REGION Network 14: Reset Manual Mode
   // Reset Manual mode when loose input flag of manual orremote enable kicks in
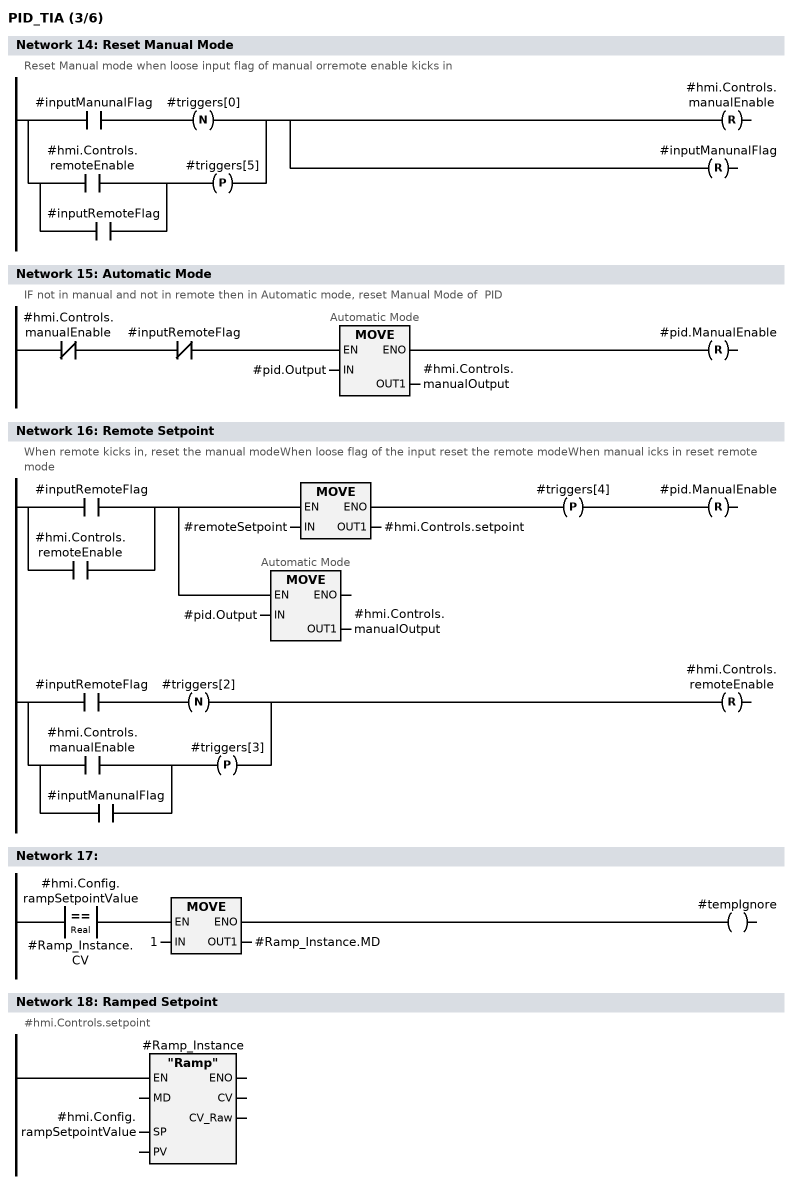
   RUNG wire#powerrail
      Contact( #inputManunalFlag )
      N_Trig( #triggers[0] )
      wire#w1
      R_Coil( #hmi.Controls.manualEnable )
   END_RUNG
   RUNG wire#powerrail
      Contact( #hmi.Controls.remoteEnable )
      wire#w2
      P_Trig( #triggers[5] )
   END_RUNG wire#w1
   RUNG wire#powerrail
      Contact( #inputRemoteFlag )
   END_RUNG wire#w2
   RUNG wire#w1
      R_Coil( #inputManunalFlag )
   END_RUNG
   // the same network as SCL:
   #_w1 := NOT #inputManunalFlag AND #triggers[0];   // falling edge
   #triggers[0] := #inputManunalFlag;
   #_w2 := #hmi.Controls.remoteEnable OR #inputRemoteFlag;
   #_w3 := #_w2 AND NOT #triggers[5];   // rising edge
   #triggers[5] := #_w2;
   IF #_w1 OR #_w3 THEN
       #hmi.Controls.manualEnable := FALSE;
       #inputManunalFlag := FALSE;
   END_IF;
END_REGION

REGION Network 15: Automatic Mode
   // IF not in manual and not in remote then in Automatic mode, reset Manual Mode of  PID
   RUNG wire#powerrail
      I_Contact( #hmi.Controls.manualEnable )
      I_Contact( #inputRemoteFlag )
      Move(in := #pid.Output, out1 => #hmi.Controls.manualOutput)   // Automatic Mode
      R_Coil( #pid.ManualEnable )
   END_RUNG
   // the same network as SCL:
   IF NOT #hmi.Controls.manualEnable AND NOT #inputRemoteFlag THEN
       #hmi.Controls.manualOutput := #pid.Output;   // Automatic Mode
       #pid.ManualEnable := FALSE;
   END_IF;
END_REGION

REGION Network 16: Remote Setpoint
   // When remote kicks in, reset the manual modeWhen loose flag of the input reset the remote modeWhen manual icks in reset remote mode
   RUNG wire#powerrail
      Contact( #inputRemoteFlag )
      wire#w1
      Move(in := #remoteSetpoint, out1 => #hmi.Controls.setpoint)
      P_Trig( #triggers[4] )
      R_Coil( #pid.ManualEnable )
   END_RUNG
   RUNG wire#powerrail
      Contact( #hmi.Controls.remoteEnable )
   END_RUNG wire#w1
   RUNG wire#w1
      Move(in := #pid.Output, out1 => #hmi.Controls.manualOutput)   // Automatic Mode
   END_RUNG
   RUNG wire#powerrail
      Contact( #inputRemoteFlag )
      N_Trig( #triggers[2] )
      wire#w2
      R_Coil( #hmi.Controls.remoteEnable )
   END_RUNG
   RUNG wire#powerrail
      Contact( #hmi.Controls.manualEnable )
      wire#w3
      P_Trig( #triggers[3] )
   END_RUNG wire#w2
   RUNG wire#powerrail
      Contact( #inputManunalFlag )
   END_RUNG wire#w3
   // the same network as SCL:
   #_w1 := #inputRemoteFlag OR #hmi.Controls.remoteEnable;
   IF #_w1 THEN #hmi.Controls.setpoint := #remoteSetpoint; END_IF;
   #_w2 := #_w1 AND NOT #triggers[4];   // rising edge
   #triggers[4] := #_w1;
   IF #_w2 THEN #pid.ManualEnable := FALSE; END_IF;
   IF #_w1 THEN
       #hmi.Controls.manualOutput := #pid.Output;   // Automatic Mode
   END_IF;
   #_w3 := NOT #inputRemoteFlag AND #triggers[2];   // falling edge
   #triggers[2] := #inputRemoteFlag;
   #_w4 := #hmi.Controls.manualEnable OR #inputManunalFlag;
   #_w5 := #_w4 AND NOT #triggers[3];   // rising edge
   #triggers[3] := #_w4;
   IF #_w3 OR #_w5 THEN #hmi.Controls.remoteEnable := FALSE; END_IF;
END_REGION

REGION Network 17
   RUNG wire#powerrail
      { S7_Templates := "SrcType := Real" } EQ_Contact(in1 := #hmi.Config.rampSetpointValue, in2 := #Ramp_Instance.CV)
      Move(in := 1, out1 => #Ramp_Instance.MD)
      Coil( #tempIgnore )
   END_RUNG
   // the same network as SCL:
   #_w1 := #hmi.Config.rampSetpointValue = #Ramp_Instance.CV;
   IF #_w1 THEN #Ramp_Instance.MD := 1; END_IF;
   #tempIgnore := #_w1;
END_REGION

REGION Network 18: Ramped Setpoint
   // #hmi.Controls.setpoint
   RUNG wire#powerrail
      #Ramp_Instance(MD :=, SP := #hmi.Config.rampSetpointValue, PV :=, CV =>, CV_Raw =>)
   END_RUNG
   // the same network as SCL:
   #Ramp_Instance(SP := #hmi.Config.rampSetpointValue);   // "Ramp"
END_REGION

REGION Network 19: Setpoint Control
   // If ramp enabled then move ramped setpointif ramp disabled then move hmi setpoint
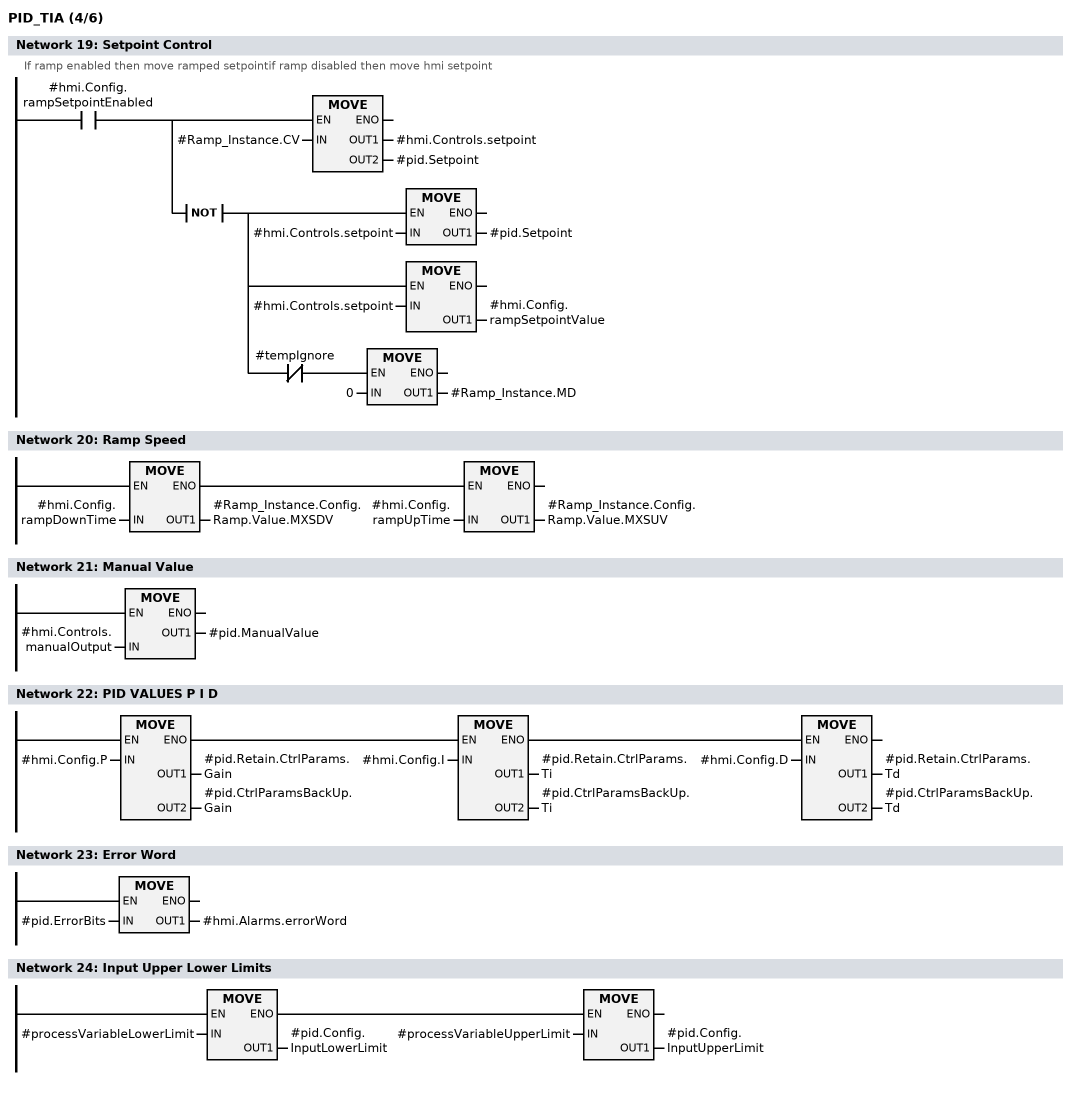
   RUNG wire#powerrail
      Contact( #hmi.Config.rampSetpointEnabled )
      wire#w1
      Move(in := #Ramp_Instance.CV, out1 => #hmi.Controls.setpoint, out2 => #pid.Setpoint)
   END_RUNG
   RUNG wire#w1
      Not()
      wire#w2
      Move(in := #hmi.Controls.setpoint, out1 => #pid.Setpoint)
   END_RUNG
   RUNG wire#w2
      Move(in := #hmi.Controls.setpoint, out1 => #hmi.Config.rampSetpointValue)
   END_RUNG
   RUNG wire#w2
      I_Contact( #tempIgnore )
      Move(in := 0, out1 => #Ramp_Instance.MD)
   END_RUNG
   // the same network as SCL:
   IF #hmi.Config.rampSetpointEnabled THEN
       #hmi.Controls.setpoint := #Ramp_Instance.CV;
       #pid.Setpoint := #Ramp_Instance.CV;
   END_IF;
   #_w1 := NOT #hmi.Config.rampSetpointEnabled;
   IF #_w1 THEN
       #pid.Setpoint := #hmi.Controls.setpoint;
       #hmi.Config.rampSetpointValue := #hmi.Controls.setpoint;
   END_IF;
   IF #_w1 AND NOT #tempIgnore THEN #Ramp_Instance.MD := 0; END_IF;
END_REGION

REGION Network 20: Ramp Speed
   RUNG wire#powerrail
      Move(in := #hmi.Config.rampDownTime, out1 => #Ramp_Instance.Config.Ramp.Value.MXSDV)
      Move(in := #hmi.Config.rampUpTime, out1 => #Ramp_Instance.Config.Ramp.Value.MXSUV)
   END_RUNG
   // the same network as SCL:
   #Ramp_Instance.Config.Ramp.Value.MXSDV := #hmi.Config.rampDownTime;
   #Ramp_Instance.Config.Ramp.Value.MXSUV := #hmi.Config.rampUpTime;
END_REGION

REGION Network 21: Manual Value
   RUNG wire#powerrail
      Move(in := #hmi.Controls.manualOutput, out1 => #pid.ManualValue)
   END_RUNG
   // the same network as SCL:
   #pid.ManualValue := #hmi.Controls.manualOutput;
END_REGION

REGION Network 22: PID VALUES P I D
   RUNG wire#powerrail
      Move(in := #hmi.Config.P, out1 => #pid.Retain.CtrlParams.Gain, out2 => #pid.CtrlParamsBackUp.Gain)
      Move(in := #hmi.Config.I, out1 => #pid.Retain.CtrlParams.Ti, out2 => #pid.CtrlParamsBackUp.Ti)
      Move(in := #hmi.Config.D, out1 => #pid.Retain.CtrlParams.Td, out2 => #pid.CtrlParamsBackUp.Td)
   END_RUNG
   // the same network as SCL:
   #pid.Retain.CtrlParams.Gain := #hmi.Config.P;
   #pid.CtrlParamsBackUp.Gain := #hmi.Config.P;
   #pid.Retain.CtrlParams.Ti := #hmi.Config.I;
   #pid.CtrlParamsBackUp.Ti := #hmi.Config.I;
   #pid.Retain.CtrlParams.Td := #hmi.Config.D;
   #pid.CtrlParamsBackUp.Td := #hmi.Config.D;
END_REGION

REGION Network 23: Error Word
   RUNG wire#powerrail
      Move(in := #pid.ErrorBits, out1 => #hmi.Alarms.errorWord)
   END_RUNG
   // the same network as SCL:
   #hmi.Alarms.errorWord := #pid.ErrorBits;
END_REGION

REGION Network 24: Input Upper Lower Limits
   RUNG wire#powerrail
      Move(in := #processVariableLowerLimit, out1 => #pid.Config.InputLowerLimit)
      Move(in := #processVariableUpperLimit, out1 => #pid.Config.InputUpperLimit)
   END_RUNG
   // the same network as SCL:
   #pid.Config.InputLowerLimit := #processVariableLowerLimit;
   #pid.Config.InputUpperLimit := #processVariableUpperLimit;
END_REGION

REGION Network 25: Input to Input PID
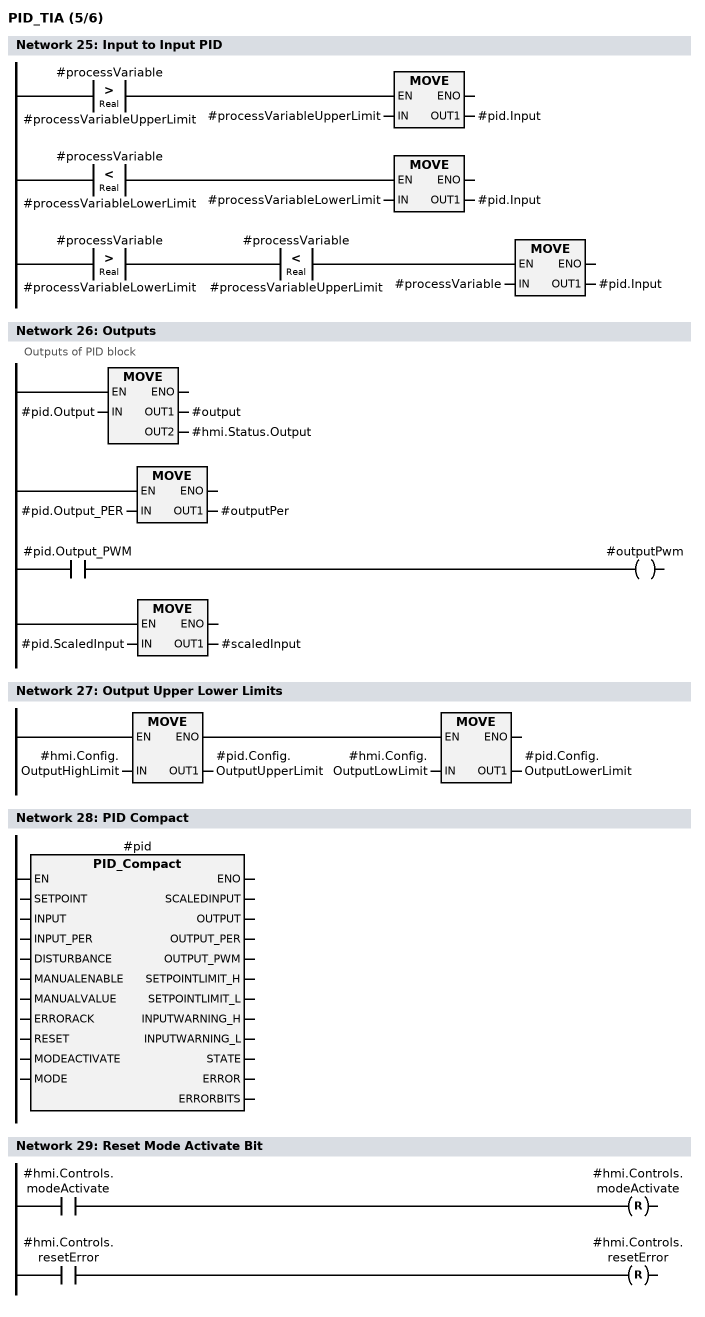
   RUNG wire#powerrail
      { S7_Templates := "SrcType := Real" } GT_Contact(in1 := #processVariable, in2 := #processVariableUpperLimit)
      Move(in := #processVariableUpperLimit, out1 => #pid.Input)
   END_RUNG
   RUNG wire#powerrail
      { S7_Templates := "SrcType := Real" } LT_Contact(in1 := #processVariable, in2 := #processVariableLowerLimit)
      Move(in := #processVariableLowerLimit, out1 => #pid.Input)
   END_RUNG
   RUNG wire#powerrail
      { S7_Templates := "SrcType := Real" } GT_Contact(in1 := #processVariable, in2 := #processVariableLowerLimit)
      { S7_Templates := "SrcType := Real" } LT_Contact(in1 := #processVariable, in2 := #processVariableUpperLimit)
      Move(in := #processVariable, out1 => #pid.Input)
   END_RUNG
   // the same network as SCL:
   IF #processVariable > #processVariableUpperLimit THEN #pid.Input := #processVariableUpperLimit; END_IF;
   IF #processVariable < #processVariableLowerLimit THEN #pid.Input := #processVariableLowerLimit; END_IF;
   IF (#processVariable > #processVariableLowerLimit) AND (#processVariable < #processVariableUpperLimit) THEN
       #pid.Input := #processVariable;
   END_IF;
END_REGION

REGION Network 26: Outputs
   // Outputs of PID block
   RUNG wire#powerrail
      Move(in := #pid.Output, out1 => #output, out2 => #hmi.Status.Output)
   END_RUNG
   RUNG wire#powerrail
      Move(in := #pid.Output_PER, out1 => #outputPer)
   END_RUNG
   RUNG wire#powerrail
      Contact( #pid.Output_PWM )
      Coil( #outputPwm )
   END_RUNG
   RUNG wire#powerrail
      Move(in := #pid.ScaledInput, out1 => #scaledInput)
   END_RUNG
   // the same network as SCL:
   #output := #pid.Output;
   #hmi.Status.Output := #pid.Output;
   #outputPer := #pid.Output_PER;
   #outputPwm := #pid.Output_PWM;
   #scaledInput := #pid.ScaledInput;
END_REGION

REGION Network 27: Output Upper Lower Limits
   RUNG wire#powerrail
      Move(in := #hmi.Config.OutputHighLimit, out1 => #pid.Config.OutputUpperLimit)
      Move(in := #hmi.Config.OutputLowLimit, out1 => #pid.Config.OutputLowerLimit)
   END_RUNG
   // the same network as SCL:
   #pid.Config.OutputUpperLimit := #hmi.Config.OutputHighLimit;
   #pid.Config.OutputLowerLimit := #hmi.Config.OutputLowLimit;
END_REGION

REGION Network 28: PID Compact
   #pid();   // PID_Compact
END_REGION

REGION Network 29: Reset Mode Activate Bit
   RUNG wire#powerrail
      Contact( #hmi.Controls.modeActivate )
      R_Coil( #hmi.Controls.modeActivate )
   END_RUNG
   RUNG wire#powerrail
      Contact( #hmi.Controls.resetError )
      R_Coil( #hmi.Controls.resetError )
   END_RUNG
   // the same network as SCL:
   IF #hmi.Controls.modeActivate THEN #hmi.Controls.modeActivate := FALSE; END_IF;
   IF #hmi.Controls.resetError THEN #hmi.Controls.resetError := FALSE; END_IF;
END_REGION

REGION Network 30: PV Tracking
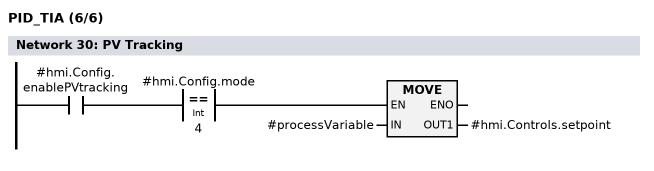
   RUNG wire#powerrail
      Contact( #hmi.Config.enablePVtracking )
      { S7_Templates := "SrcType := Int" } EQ_Contact(in1 := #hmi.Config.mode, in2 := 4)
      Move(in := #processVariable, out1 => #hmi.Controls.setpoint)
   END_RUNG
   // the same network as SCL:
   IF #hmi.Config.enablePVtracking AND (#hmi.Config.mode = 4) THEN
       #hmi.Controls.setpoint := #processVariable;
   END_IF;
END_REGION
END_FUNCTION_BLOCK

// folder: 1}Library/Pumps

FUNCTION_BLOCK "SimpleMotorStater"   // FB823, LAD
{ S7_Optimized_Access := 'TRUE' }
VERSION : 0.1
   VAR_INPUT
      OP_Mode : Bool;   // Output Mode for the Stop CMD if True( Normal Open Output) If False ( Normal Close Output)
      ON : Bool;   // Motor On
      OFF : Bool := TRUE;   // Motor OFF
      CF : Bool;   // Status- Contact Feedback
      IL : Bool := TRUE;   // status-Interlock
      "Lead Control" : Bool := TRUE;
   END_VAR
   VAR_OUTPUT
      Stop_CMD : Bool := TRUE;   // Stop Command for the Motor
      Start_CMD : Bool;   // Start Command for the Motor
      RST : Bool;   // Reset Overload
   END_VAR
   VAR
      HMI : Struct   // Data Struct for HMI
         Controls : Struct
            Start : Bool;
            Stop : Bool := TRUE;
            Reset : Bool;
            Lockout : Bool;
         END_STRUCT;
         Status : Struct
            Mode : Bool;   // Output Mode for the Stop CMD if True Normal Open Output (NO) If False Normal Close Output (NC)
            CF : Bool;   // Status- Contact Feedback
            IL : Bool;   // Status-Interlock
            State : Int;   // 0=off, 1=on, 2=fault,3= Lockout
         END_STRUCT;
      END_STRUCT;
   END_VAR
   VAR RETAIN
      Config : Struct
         HMI : Struct
            Start_PT : Time := T#500MS;   // Start CMD Pulse Time
            Stop_PT : Time := T#500MS;   // Stop CMD Pulse Time
            CF_Delay : Time := T#10s;   // Contact Feedback Delay Time
            NCresetDelay : Time := T#1s;   // time to Set stop on went in NC Mode
            Enable_HMI_Controls : Int;   // MODE 1 PLC CTRL / MODE 2 HMII
         END_STRUCT;
      END_STRUCT;
   END_VAR
   VAR
      OS : Struct
         ON : Bool;
         OFF : Bool;
         HMION : Bool;
         HMIOFF : Bool;
         CF_PULSE : Bool;
         ILPOS : Bool;
         PULSE : Bool;
      END_STRUCT;
      STOP_CMD_TOF : TOF_TIME;   // Stop CMD Pulse Timer
      START_CMD_TOF : TOF_TIME;   // Start CMD Pulse Timer
      CF_Delay_TON : TOF_TIME;   // Contact Feedback Delay Timer
      DelayforReset : TON_TIME;
      FaultTimer : IEC_TIMER;
      Fault : Bool;
      "Lockout Trig" : Bool;
   END_VAR
   VAR_TEMP
      STOP : Bool;
   END_VAR
   VAR_TEMP   // added for the SCL form of the ladder/FBD networks
      _w1 : Bool;
      _w2 : Bool;
      _w3 : Bool;
      _w4 : Bool;
      _w5 : Bool;
      _w6 : Bool;
      _w7 : Bool;
      _w8 : Bool;
   END_VAR
BEGIN

REGION Network 1: Status-Interlock
   // Interloack Status for HMI
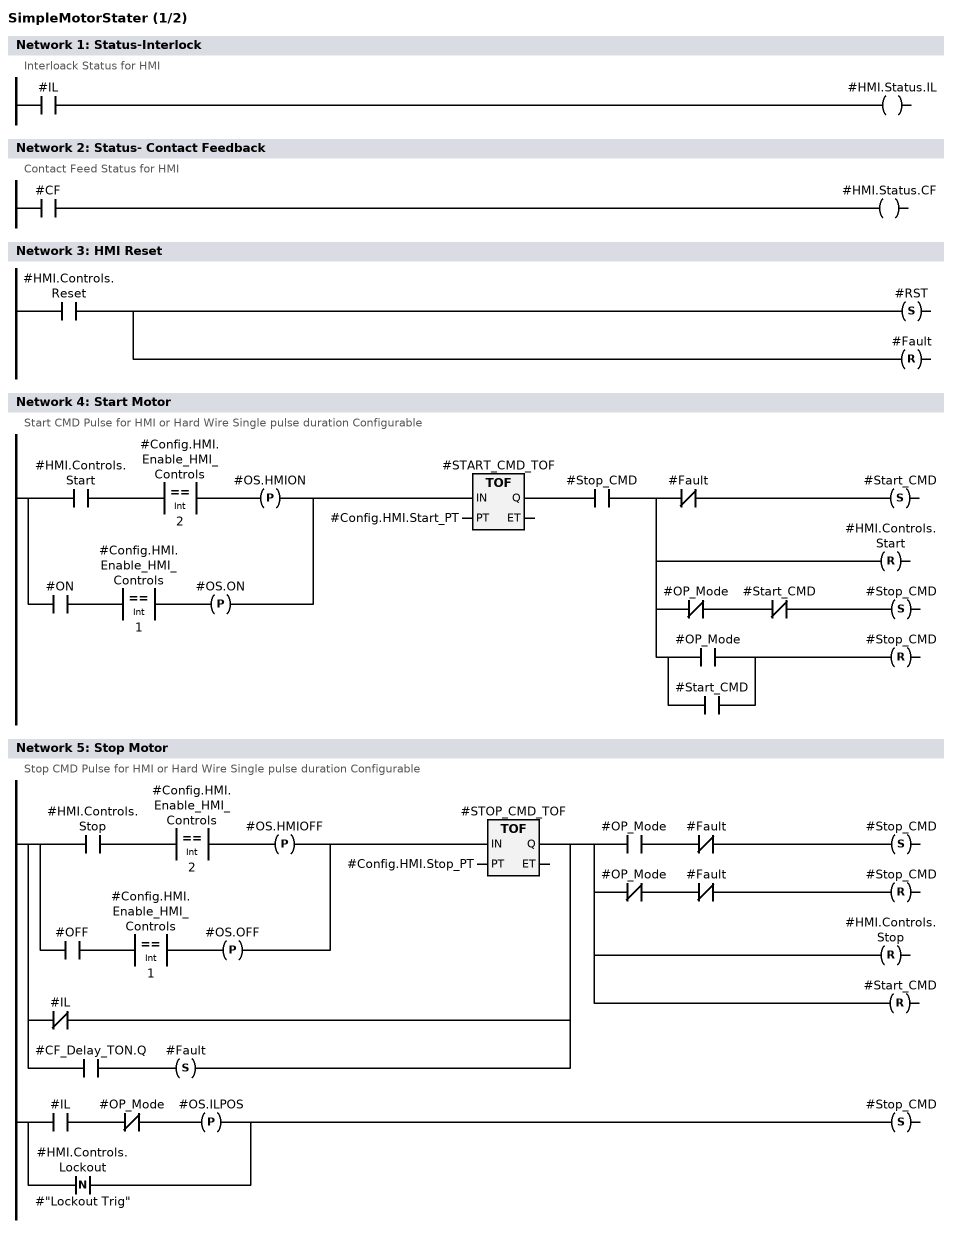
   RUNG wire#powerrail
      Contact( #IL )
      Coil( #HMI.Status.IL )
   END_RUNG
   // the same network as SCL:
   #HMI.Status.IL := #IL;
END_REGION

REGION Network 2: Status- Contact Feedback
   // Contact Feed Status for HMI
   RUNG wire#powerrail
      Contact( #CF )
      Coil( #HMI.Status.CF )
   END_RUNG
   // the same network as SCL:
   #HMI.Status.CF := #CF;
END_REGION

REGION Network 3: HMI Reset
   RUNG wire#powerrail
      Contact( #HMI.Controls.Reset )
      wire#w1
      S_Coil( #RST )
   END_RUNG
   RUNG wire#w1
      R_Coil( #Fault )
   END_RUNG
   // the same network as SCL:
   IF #HMI.Controls.Reset THEN
       #RST := TRUE;
       #Fault := FALSE;
   END_IF;
END_REGION

REGION Network 4: Start Motor
   // Start CMD Pulse for HMI or Hard Wire Single pulse duration Configurable
   #_w1 := #HMI.Controls.Start AND (#Config.HMI.Enable_HMI_Controls = 2);
   #_w2 := #_w1 AND NOT #OS.HMION;   // rising edge
   #OS.HMION := #_w1;
   #_w3 := #ON AND (#Config.HMI.Enable_HMI_Controls = 1);
   #_w4 := #_w3 AND NOT #OS.ON;   // rising edge
   #OS.ON := #_w3;
   #START_CMD_TOF(IN := #_w2 OR #_w4, PT := #Config.HMI.Start_PT);   // TOF
   #_w5 := #START_CMD_TOF.Q AND #Stop_CMD;
   IF #_w5 AND NOT #Fault THEN #Start_CMD := TRUE; END_IF;
   IF #_w5 THEN #HMI.Controls.Start := FALSE; END_IF;
   IF #_w5 AND NOT #OP_Mode AND NOT #Start_CMD THEN #Stop_CMD := TRUE; END_IF;
   IF #_w5 AND (#OP_Mode OR #Start_CMD) THEN #Stop_CMD := FALSE; END_IF;
END_REGION

REGION Network 5: Stop Motor
   // Stop CMD Pulse for HMI or Hard Wire Single pulse duration Configurable
   #_w1 := #HMI.Controls.Stop AND (#Config.HMI.Enable_HMI_Controls = 2);
   #_w2 := #_w1 AND NOT #OS.HMIOFF;   // rising edge
   #OS.HMIOFF := #_w1;
   #_w3 := #OFF AND (#Config.HMI.Enable_HMI_Controls = 1);
   #_w4 := #_w3 AND NOT #OS.OFF;   // rising edge
   #OS.OFF := #_w3;
   #STOP_CMD_TOF(IN := #_w2 OR #_w4, PT := #Config.HMI.Stop_PT);   // TOF
   IF #CF_Delay_TON.Q THEN #Fault := TRUE; END_IF;
   #_w5 := #STOP_CMD_TOF.Q OR NOT #IL OR #CF_Delay_TON.Q;
   IF #_w5 AND #OP_Mode AND NOT #Fault THEN #Stop_CMD := TRUE; END_IF;
   IF #_w5 AND NOT #OP_Mode AND NOT #Fault THEN #Stop_CMD := FALSE; END_IF;
   IF #_w5 THEN
       #HMI.Controls.Stop := FALSE;
       #Start_CMD := FALSE;
   END_IF;
   #_w6 := #IL AND NOT #OP_Mode;
   #_w7 := #_w6 AND NOT #OS.ILPOS;   // rising edge
   #OS.ILPOS := #_w6;
   #_w8 := NOT #HMI.Controls.Lockout AND #"Lockout Trig";   // falling edge of #HMI.Controls.Lockout
   #"Lockout Trig" := #HMI.Controls.Lockout;
   IF #_w7 OR #_w8 THEN #Stop_CMD := TRUE; END_IF;
END_REGION

REGION Network 6: Delay for Contact feedback
   // Timer Delay for For Feedback Duration Configurable
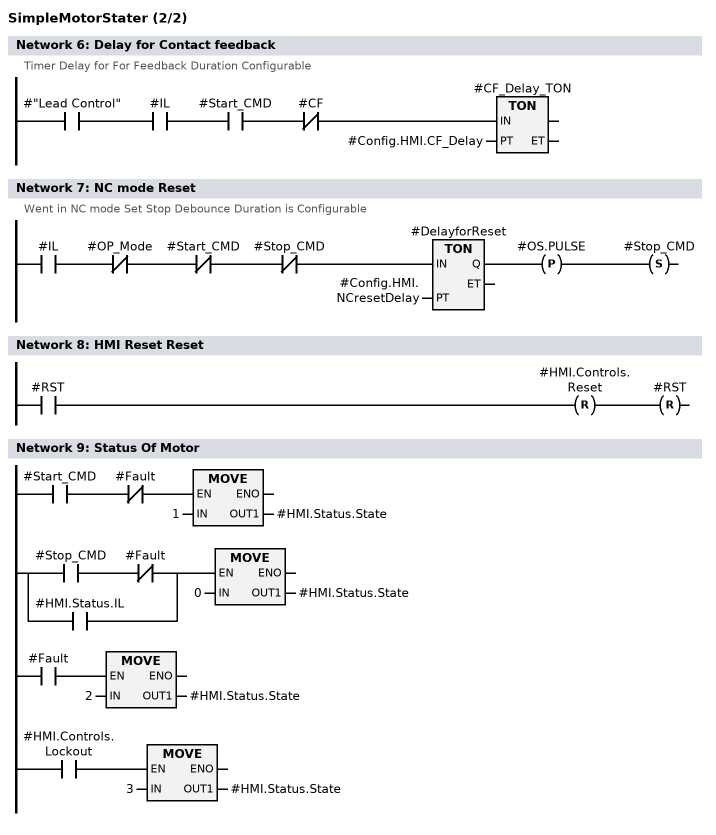
   #CF_Delay_TON(IN := #"Lead Control" AND #IL AND #Start_CMD AND NOT #CF, PT := #Config.HMI.CF_Delay);   // TON
END_REGION

REGION Network 7: NC mode Reset
   // Went in NC mode Set Stop Debounce Duration is Configurable
   #DelayforReset(IN := #IL AND NOT #OP_Mode AND NOT #Start_CMD AND NOT #Stop_CMD,   // TON
                  PT := #Config.HMI.NCresetDelay);
   #_w1 := #DelayforReset.Q AND NOT #OS.PULSE;   // rising edge
   #OS.PULSE := #DelayforReset.Q;
   IF #_w1 THEN #Stop_CMD := TRUE; END_IF;
END_REGION

REGION Network 8: HMI Reset Reset
   RUNG wire#powerrail
      Contact( #RST )
      R_Coil( #HMI.Controls.Reset )
      R_Coil( #RST )
   END_RUNG
   // the same network as SCL:
   IF #RST THEN
       #HMI.Controls.Reset := FALSE;
       #RST := FALSE;
   END_IF;
END_REGION

REGION Network 9: Status Of Motor
   RUNG wire#powerrail
      Contact( #Start_CMD )
      I_Contact( #Fault )
      Move(in := 1, out1 => #HMI.Status.State)
   END_RUNG
   RUNG wire#powerrail
      Contact( #Stop_CMD )
      I_Contact( #Fault )
      wire#w1
      Move(in := 0, out1 => #HMI.Status.State)
   END_RUNG
   RUNG wire#powerrail
      Contact( #HMI.Status.IL )
   END_RUNG wire#w1
   RUNG wire#powerrail
      Contact( #Fault )
      Move(in := 2, out1 => #HMI.Status.State)
   END_RUNG
   RUNG wire#powerrail
      Contact( #HMI.Controls.Lockout )
      Move(in := 3, out1 => #HMI.Status.State)
   END_RUNG
   // the same network as SCL:
   IF #Start_CMD AND NOT #Fault THEN #HMI.Status.State := 1; END_IF;
   IF (#Stop_CMD AND NOT #Fault) OR #HMI.Status.IL THEN #HMI.Status.State := 0; END_IF;
   IF #Fault THEN #HMI.Status.State := 2; END_IF;
   IF #HMI.Controls.Lockout THEN #HMI.Status.State := 3; END_IF;
END_REGION
END_FUNCTION_BLOCK

// folder: 1}Library/Ramp

FUNCTION_BLOCK "Ramp_v2"   // FB4, SCL
{ S7_Optimized_Access := 'TRUE' }
VERSION : 0.1
   VAR
      Enable : Bool;   // Enable the Block
      Parameters : Struct
         End_SP : Real;   // End Setpoint
         Working_SP : Real;   // Working Setpoint
         PV : Real;   // Process Value
         Rate : Int := 3;   // Ramp Rate
         RateTime : Time := T#1m;
         MaxRate : Int := 10;   // Max Ramp Rate
      END_STRUCT;
      FirstCycle : Bool;   // First Cycle after enable the block
      TimeSlide : DInt;
      TimeSP : Time;
      "Time" : IEC_TIMER;
      Control : Struct
         OS : Bool;
         CountUp : Bool;
         RampDone : Bool;
      END_STRUCT;
   END_VAR
   VAR CONSTANT
      AddValue : Real := 0.1;   // Value to add to the Working SP within the Rate
      Time0 : Time;
   END_VAR
BEGIN
   //Ramp SP Block
   //

   IF #Enable THEN     //Enable the execution of the block

       IF #Parameters.Rate > #Parameters.MaxRate THEN    //Rate should not be greater that maxRate

           #Parameters.Rate := #Parameters.MaxRate;      //if Rate is greater that maxRate then Rate iqual to maxRate.

       END_IF;

       IF #Parameters.PV > 0.0 THEN   //Process Value greater that 0.0
           //First Cycle after enable the block and PV greater that 0.0
           IF #FirstCycle THEN
               #FirstCycle := False;
               #Parameters.Working_SP := #Parameters.PV;     //Start Controlling from the Process Value (PV).
               #Control.OS := TRUE;
           END_IF;
       END_IF;

       #TimeSlide := TIME_TO_DINT(#Parameters.RateTime);   //Convert Rate time to Dint data type
       #TimeSlide := #TimeSlide / #Parameters.Rate;        //get the time to do the increase of the Working SP 
       #TimeSP := DINT_TO_TIME(#TimeSlide);                //Convert the time increase to a time data time

       #Control.CountUp := #Time.Q AND #TimeSP > #Time0;

       IF #Control.CountUp  THEN
           #Parameters.Working_SP:=#Parameters.Working_SP+1;
       END_IF;

       IF #Parameters.Working_SP >= #Parameters.End_SP THEN
           #Parameters.Working_SP := #Parameters.End_SP;
           #Control.RampDone := TRUE;
       ELSE
           #Control.RampDone := FALSE;
       END_IF;
   ELSE
       #FirstCycle := TRUE;
       #Control.OS := FALSE;
       #Parameters.Working_SP := 0.0;

   END_IF;

   #Time.TON(IN := #Control.OS AND NOT #Control.CountUp AND NOT #Control.RampDone,
             PT := #TimeSP);
END_FUNCTION_BLOCK

FUNCTION_BLOCK "Ramp"   // FB701, LAD
{ S7_Optimized_Access := 'FALSE' }
VERSION : 1.0
   VAR_INPUT
      MD : Int := 1;   // FB Mode "0=No Ramp" "1=Ramp"
      SP : Real;   // Setpoint
      PV : Real;   // Process Value
   END_VAR
   VAR_OUTPUT
      CV : Real;   // Control Value in Real Data Type
      CV_Raw : Int;   // Control Value in INT Data Type
   END_VAR
   VAR
      Control : Struct
         SP : Real;   // Current SP / Can be configurable in HMI if SIM is enabled
         Hold : Bool;   // Hold last commanded CV
      END_STRUCT;
      Config : Struct
         Unscale : Struct
            HL : Real := 100.0;   // Unscale High Limit
            LL : Real;   // Unscale Low Limit
            Bipolar : Bool;   // Enable/Disable Bipolar Value
         END_STRUCT;
         Ramp : Struct
            PT : Struct   // Preset Time
               Up : Time := T#100ms;   // Ramp Up Preset Time
               Down : Time := T#100ms;   // Ramp Down Preset Time
            END_STRUCT;
            Value : Struct
               MXSUV : Real := 1.0;   // Max Step/Ramp Up Value
               MXSDV : Real := 1.0;   // Max Step/Ramp Down Value
            END_STRUCT;
         END_STRUCT;
         Deadband : Struct
            UDW : Real := 0.5;   // Upper Deadband Width
            LDW : Real := 0.5;   // Lower Deadband Width
         END_STRUCT;
         TPV : Bool;   // Enable Process Variable Tracking
         SIM : Bool;   // Simulate SP
      END_STRUCT;
      Status : Struct
         USRV : Word;   // Unscale RET_VAL
         PV : Real;   // Current Process Value
         CV : Real;   // Current Control Value
      END_STRUCT;
      Oneshot : Struct
         Up : Bool;
         Down : Bool;
      END_STRUCT;
      RUIT : TON_TIME;   // Ramp Up Interval Time
      RDIT : TON_TIME;   // Ramp Down Interval Time
      Deviation : "Deviation";
   END_VAR
   VAR_TEMP
      PVHL : Real;   // PV High Limit when tracking is enabled
      PVLL : Real;   // PV Low Limit when tracking is enabled
   END_VAR
   VAR_TEMP   // added for the SCL form of the ladder/FBD networks
      _w1 : Bool;
   END_VAR
BEGIN

REGION Network 1: Enablee/Disable SP Simulation
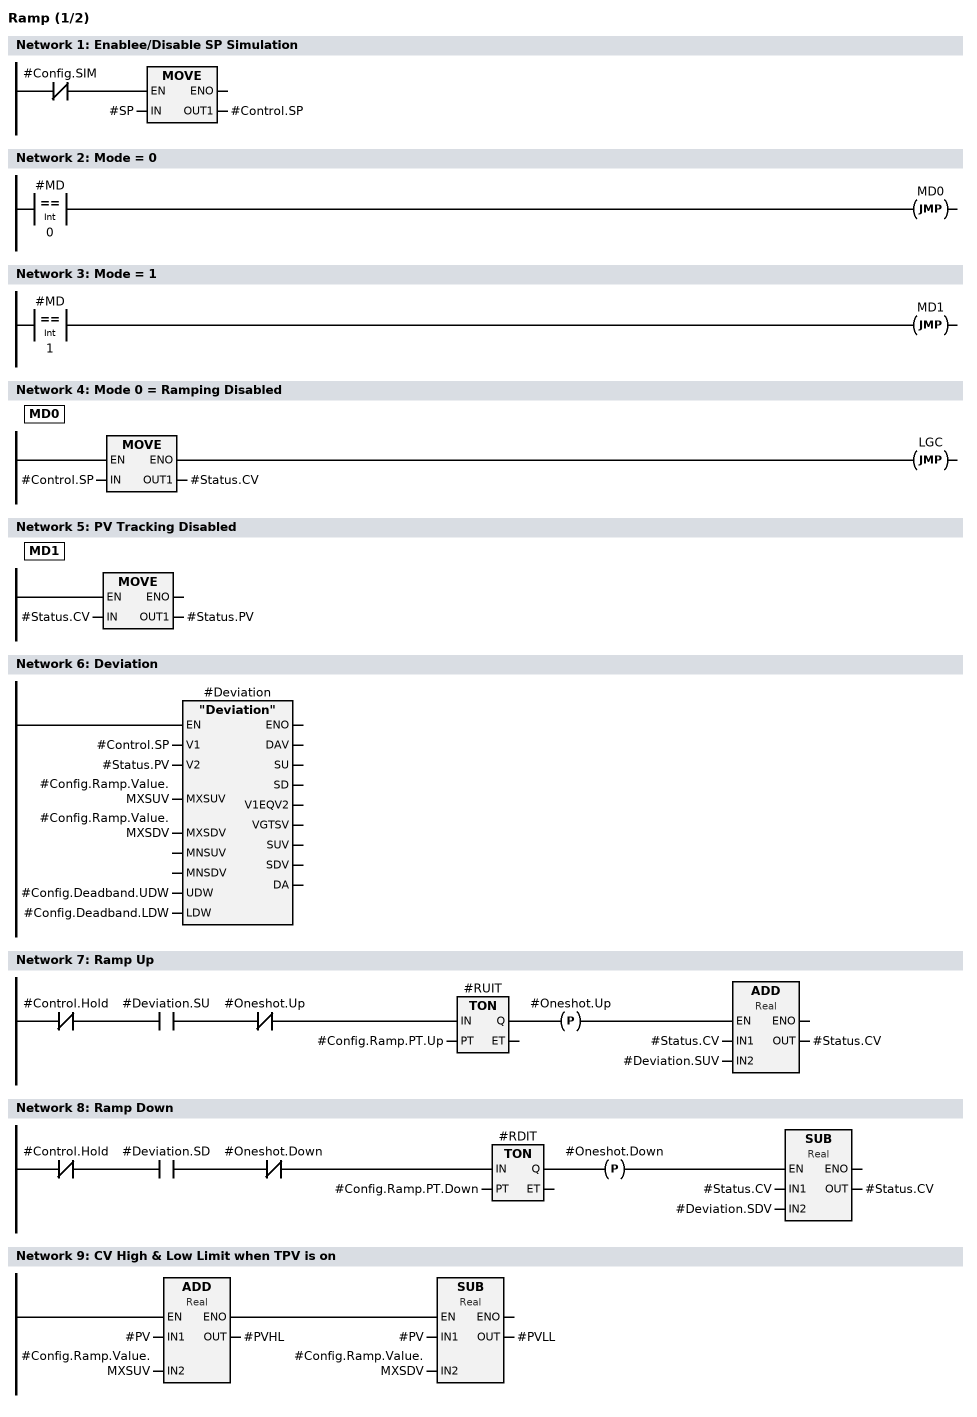
   RUNG wire#powerrail
      I_Contact( #Config.SIM )
      { S7_GenerateENO := "TRUE" } Move(in := #SP, out1 => #Control.SP)
   END_RUNG
   // the same network as SCL:
   IF NOT #Config.SIM THEN #Control.SP := #SP; END_IF;
END_REGION

REGION Network 2: Mode = 0
   RUNG wire#powerrail
      { S7_Templates := "SrcType := Int" } EQ_Contact(in1 := #MD, in2 := 0)
      JumpCoil( MD0 )
   END_RUNG
   // the same network as SCL:
   IF #MD = 0 THEN GOTO MD0; END_IF;
END_REGION

REGION Network 3: Mode = 1
   RUNG wire#powerrail
      { S7_Templates := "SrcType := Int" } EQ_Contact(in1 := #MD, in2 := 1)
      JumpCoil( MD1 )
   END_RUNG
   // the same network as SCL:
   IF #MD = 1 THEN GOTO MD1; END_IF;
END_REGION

REGION Network 4: Mode 0 = Ramping Disabled
   Label( MD0 )
   RUNG wire#powerrail
      { S7_GenerateENO := "TRUE" } Move(in := #Control.SP, out1 => #Status.CV)
      JumpCoil( LGC )
   END_RUNG
   // the same network as SCL:
   // ENO of a box is taken as its EN; it also drops when the box reports an error
   MD0:
   #Status.CV := #Control.SP;
   GOTO LGC;
END_REGION

REGION Network 5: PV Tracking Disabled
   Label( MD1 )
   RUNG wire#powerrail
      { S7_GenerateENO := "TRUE" } Move(in := #Status.CV, out1 => #Status.PV)
   END_RUNG
   // the same network as SCL:
   MD1:
   #Status.PV := #Status.CV;
END_REGION

REGION Network 6: Deviation
   RUNG wire#powerrail
      #Deviation(V1 := #Control.SP, V2 := #Status.PV, MXSUV := #Config.Ramp.Value.MXSUV, MXSDV := #Config.Ramp.Value.MXSDV, MNSUV :=, MNSDV :=, UDW := #Config.Deadband.UDW, LDW := #Config.Deadband.LDW, DAV =>, SU =>, SD =>, V1EQV2 =>, VGTSV =>, SUV =>, SDV =>, DA =>)
   END_RUNG
   // the same network as SCL:
   #Deviation(V1 := #Control.SP,   // "Deviation"
              V2 := #Status.PV,
              MXSUV := #Config.Ramp.Value.MXSUV,
              MXSDV := #Config.Ramp.Value.MXSDV,
              UDW := #Config.Deadband.UDW,
              LDW := #Config.Deadband.LDW);
END_REGION

REGION Network 7: Ramp Up
   #RUIT(IN := NOT #Control.Hold AND #Deviation.SU AND NOT #Oneshot.Up, PT := #Config.Ramp.PT.Up);   // TON
   #_w1 := #RUIT.Q AND NOT #Oneshot.Up;   // rising edge
   #Oneshot.Up := #RUIT.Q;
   IF #_w1 THEN #Status.CV := #Status.CV + #Deviation.SUV; END_IF;
END_REGION

REGION Network 8: Ramp Down
   #RDIT(IN := NOT #Control.Hold AND #Deviation.SD AND NOT #Oneshot.Down, PT := #Config.Ramp.PT.Down);   // TON
   #_w1 := #RDIT.Q AND NOT #Oneshot.Down;   // rising edge
   #Oneshot.Down := #RDIT.Q;
   IF #_w1 THEN #Status.CV := #Status.CV - #Deviation.SDV; END_IF;
END_REGION

REGION Network 9: CV High & Low Limit when TPV is on
   RUNG wire#powerrail
      { S7_Templates := "SrcType := Real"; S7_GenerateENO := "TRUE" } Add(in1 := #PV, in2 := #Config.Ramp.Value.MXSUV, out => #PVHL)
      { S7_Templates := "SrcType := Real"; S7_GenerateENO := "TRUE" } Sub(in1 := #PV, in2 := #Config.Ramp.Value.MXSDV, out => #PVLL)
   END_RUNG
   // the same network as SCL:
   // ENO of a box is taken as its EN; it also drops when the box reports an error
   #PVHL := #PV + #Config.Ramp.Value.MXSUV;
   #PVLL := #PV - #Config.Ramp.Value.MXSDV;
END_REGION

REGION Network 10: CV Limits when TPV is on
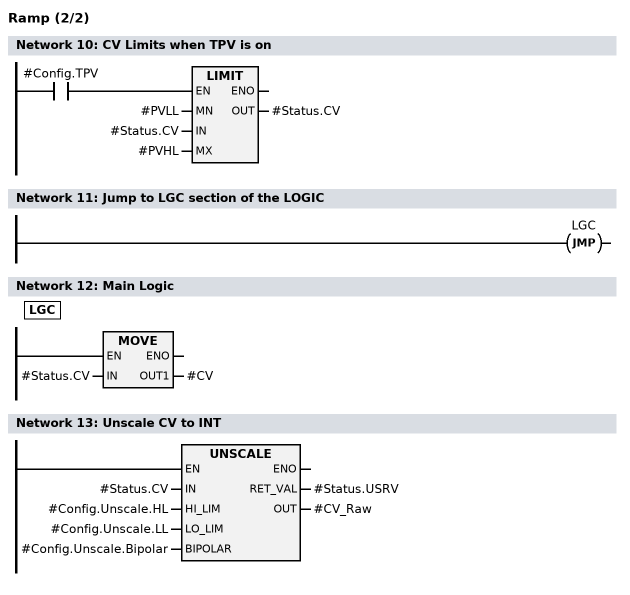
   IF #Config.TPV THEN #Status.CV := LIMIT(MN := #PVLL, IN := #Status.CV, MX := #PVHL); END_IF;
END_REGION

REGION Network 11: Jump to LGC section of the LOGIC
   RUNG wire#powerrail
      JumpCoil( LGC )
   END_RUNG
   // the same network as SCL:
   GOTO LGC;
END_REGION

REGION Network 12: Main Logic
   Label( LGC )
   RUNG wire#powerrail
      { S7_GenerateENO := "TRUE" } Move(in := #Status.CV, out1 => #CV)
   END_RUNG
   // the same network as SCL:
   LGC:
   #CV := #Status.CV;
END_REGION

REGION Network 13: Unscale CV to INT
   #Status.USRV := UNSCALE(IN := #Status.CV,
                           HI_LIM := #Config.Unscale.HL,
                           LO_LIM := #Config.Unscale.LL,
                           BIPOLAR := #Config.Unscale.Bipolar,
                           OUT => #CV_Raw);
END_REGION
END_FUNCTION_BLOCK

// folder: 1}Library/SEL Block

FUNCTION_BLOCK "LSEL"   // FB6969, LAD
{ S7_Optimized_Access := 'TRUE' }
VERSION : 0.1
   VAR_INPUT
      impulse : Bool;
   END_VAR
   VAR_OUTPUT
      done : Bool;
      busy : Bool;
      error : Bool;
      status : Word;
      frame : DWord;
      reset : Bool;
   END_VAR
   VAR
      statImpulseOld : Bool;
      HMI : Struct
         deviceName : String := 'SEL1200';
         stateCOM : Bool := TRUE;
         stateDipSwitchTD1 : Bool;
         stateDipSwitchTD2 : Bool;
         stateOutput1 : Int;   // 0=switched-off automatical, no reset possible; 1=switched-off automatical, reset possible; 2= switched-off manual; 3=switched on; 4=defect; 5=device overtemperature; 6=overload; 7=current > nominal value
         stateOutput2 : Int;   // 0=switched-off automatical, no reset possible; 1=switched-off automatical, reset possible; 2= switched-off manual; 3=switched on; 4=defect; 5=device overtemperature; 6=overload; 7=current > nominal value
         stateOutput3 : Int;   // 0=switched-off automatical, no reset possible; 1=switched-off automatical, reset possible; 2= switched-off manual; 3=switched on; 4=defect; 5=device overtemperature; 6=overload; 7=current > nominal value
         stateOutput4 : Int;   // 0=switched-off automatical, no reset possible; 1=switched-off automatical, reset possible; 2= switched-off manual; 3=switched on; 4=defect; 5=device overtemperature; 6=overload; 7=current > nominal value
         stateOutput5 : Int;   // 0=switched-off automatical, no reset possible; 1=switched-off automatical, reset possible; 2= switched-off manual; 3=switched on; 4=defect; 5=device overtemperature; 6=overload; 7=current > nominal value
         stateOutput6 : Int;   // 0=switched-off automatical, no reset possible; 1=switched-off automatical, reset possible; 2= switched-off manual; 3=switched on; 4=defect; 5=device overtemperature; 6=overload; 7=current > nominal value
         stateOutput7 : Int;   // 0=switched-off automatical, no reset possible; 1=switched-off automatical, reset possible; 2= switched-off manual; 3=switched on; 4=defect; 5=device overtemperature; 6=overload; 7=current > nominal value
         stateOutput8 : Int;   // 0=switched-off automatical, no reset possible; 1=switched-off automatical, reset possible; 2= switched-off manual; 3=switched on; 4=defect; 5=device overtemperature; 6=overload; 7=current > nominal value
         outputCurrent1 : Int;   // output current output1
         outputCurrent2 : Int;   // output current output2
         outputCurrent3 : Int;   // output current output3
         outputCurrent4 : Int;   // output current output4
         outputCurrent5 : Int;   // output current output5
         outputCurrent6 : Int;   // output current output6
         outputCurrent7 : Int;   // output current output7
         outputCurrent8 : Int;   // output current output8
         outputCurrentLimit1 : Int;   // output current limit output1
         outputCurrentLimit2 : Int;   // output current limit output2
         outputCurrentLimit3 : Int;   // output current limit output3
         outputCurrentLimit4 : Int;   // output current limit output4
         outputCurrentLimit5 : Int;   // output current limit output5
         outputCurrentLimit6 : Int;   // output current limit output6
         outputCurrentLimit7 : Int;   // output current limit output7
         outputCurrentLimit8 : Int;   // output current limit output8
         reasonOutputSwitchedOff1 : Int := 0;   // 0=output current>limit and output current<1,5xlimit for more than 5sec; 1=current output>1,5xlimit; 2=total overload; 3=Uin<19,4V and output current>limit; 4=Uin<15V; 5=Uin>30V; 6=device overtemperature; 8 to 14=Reserve; 15=default (no automatically switched off)
         reasonOutputSwitchedOff2 : Int := 0;   // 0=output current>limit and output current<1,5xlimit for more than 5sec; 1=current output>1,5xlimit; 2=total overload; 3=Uin<19,4V and output current>limit; 4=Uin<15V; 5=Uin>30V; 6=device overtemperature; 8 to 14=Reserve; 15=default (no automatically switched off)
         reasonOutputSwitchedOff3 : Int := 0;   // 0=output current>limit and output current<1,5xlimit for more than 5sec; 1=current output>1,5xlimit; 2=total overload; 3=Uin<19,4V and output current>limit; 4=Uin<15V; 5=Uin>30V; 6=device overtemperature; 8 to 14=Reserve; 15=default (no automatically switched off)
         reasonOutputSwitchedOff4 : Int := 0;   // 0=output current>limit and output current<1,5xlimit for more than 5sec; 1=current output>1,5xlimit; 2=total overload; 3=Uin<19,4V and output current>limit; 4=Uin<15V; 5=Uin>30V; 6=device overtemperature; 8 to 14=Reserve; 15=default (no automatically switched off)
         reasonOutputSwitchedOff5 : Int := 0;   // 0=output current>limit and output current<1,5xlimit for more than 5sec; 1=current output>1,5xlimit; 2=total overload; 3=Uin<19,4V and output current>limit; 4=Uin<15V; 5=Uin>30V; 6=device overtemperature; 8 to 14=Reserve; 15=default (no automatically switched off)
         reasonOutputSwitchedOff6 : Int := 0;   // 0=output current>limit and output current<1,5xlimit for more than 5sec; 1=current output>1,5xlimit; 2=total overload; 3=Uin<19,4V and output current>limit; 4=Uin<15V; 5=Uin>30V; 6=device overtemperature; 8 to 14=Reserve; 15=default (no automatically switched off)
         reasonOutputSwitchedOff7 : Int := 0;   // 0=output current>limit and output current<1,5xlimit for more than 5sec; 1=current output>1,5xlimit; 2=total overload; 3=Uin<19,4V and output current>limit; 4=Uin<15V; 5=Uin>30V; 6=device overtemperature; 8 to 14=Reserve; 15=default (no automatically switched off)
         reasonOutputSwitchedOff8 : Int := 0;   // 0=output current>limit and output current<1,5xlimit for more than 5sec; 1=current output>1,5xlimit; 2=total overload; 3=Uin<19,4V and output current>limit; 4=Uin<15V; 5=Uin>30V; 6=device overtemperature; 8 to 14=Reserve; 15=default (no automatically switched off)
         nominalOutputCurrent : Int := 3;   // nominal output current
         outputNumber : Int := 4;   // number of outputs (4 or 8)
         productState : Int := 1;   // product state
         firmwareVersion : Int := 1;   // frimware version
         startup : Int;   // 0=load dependent startup; 1=startup time tag 25ms; 2=startup time tag 200ms; 3=startup time tag 500ms
         setReset : Bool;
         stateReset : Bool;
         stateNoCommunication : Bool;
         articleNumber : String := '6EP4437-7FB00-0CX0';   // article number
         serialNumber : String := 'Q6/L1';   // serial number
      END_STRUCT;
      statTimeSave : Struct
         posEdge : DTL;
         negEdge : DTL;
         deltaTimePause : Time;
         deltaTimePauseSave : Time;
         deltaTimeImpulse : Time;
         timeIpulse : Time;
         timePause : Time;
         timeFrame : Time;
         sysTime : DTL;
         sysTimeOld : DTL;
         deltaSysTime : Time;
      END_STRUCT;
      statPosEdgeDetected : Bool;
      statPosEdgeDetectedTrigger : Bool;
      statNegEdgeDetected : Bool;
      statNegEdgeDetectedTrigger : Bool;
      statEdgeCtrl : Int;
      statArrayImpulse : Array[0..63] of Time;
      statArrayPause : Array[0..63] of Time;
      statArrayBits : Array[0..31] of Bool;
      statCntImpulse : Int;
      statCntPause : Int;
      statCntBits : Int;
      statFrame : DWord;
      statFrameOld : DWord;
      statBusy : Bool;
      statDone : Bool;
      statError : Bool;
      statErrorInt : Bool;
      statStatus : Word;
      statStatusInt : Word;
      statStateIndex : Int;
      statPauseDetected : Bool;
      statImpulseDetected : Bool;
      statIndexImpulse : Int;
      statIndexResetImpulse : Int;
      statIndexPause : Int;
      statIndexResetPause : Int;
      statIndexAddTime : Int;
      statFrameEvaluationStopp : Bool;
      statNoEvaluation : Bool;
      statStartTimerWait : Bool;
      statStartTimerSys : Bool;
      statStartWatchDogTimerPos : Bool;
      statStartWatchDogTimerNeg : Bool;
      statCycleTimeNotOk : Bool;
      instTimerWait : TON_TIME;
      instSysTimer : TON_TIME;
      instWatchDogTimerPos : TON_TIME;
      instWatchDogTimerNeg : TON_TIME;
      statDeviceName : Byte;
      statFrameID : Byte;
      statStateOutput1 : Byte;
      statStateOutput2 : Byte;
      statStateOutput3 : Byte;
      statStateOutput4 : Byte;
      statStateOutput5 : Byte;
      statStateOutput6 : Byte;
      statStateOutput7 : Byte;
      statStateOutput8 : Byte;
      statStateDipSwitchTD : Byte;
      statMeasurementsChannels : Byte;
      statOutputCurrent1 : Byte;
      statOutputCurrent2 : Byte;
      statOutputCurrent3 : Byte;
      statOutputCurrent4 : Byte;
      statOutputCurrent5 : Byte;
      statOutputCurrent6 : Byte;
      statOutputCurrent7 : Byte;
      statOutputCurrent8 : Byte;
      statOutputCurrentLimit1 : Byte;
      statOutputCurrentLimit2 : Byte;
      statOutputCurrentLimit3 : Byte;
      statOutputCurrentLimit4 : Byte;
      statOutputCurrentLimit5 : Byte;
      statOutputCurrentLimit6 : Byte;
      statOutputCurrentLimit7 : Byte;
      statOutputCurrentLimit8 : Byte;
      statNominalOutputCurrent : Byte;
      statConstructionYearByte : Byte;
      statConstructionYearChar : Char;
      statConstructionYear : Int;
      statConstructionMonthByte : Byte;
      statConstructionMonthChar : Char;
      statConstructionMonth : Int;
      statProductState : Byte;
      statFirmwareVersion : Byte;
      statVarianten11 : Byte;
      statInnovationen : Byte;
      statChannelNumber : Byte;
      statPower : Int;
      statLacquered : Bool;
      statFabricationPlace : Bool;
      statDeviceType : Bool;
      statStateInputVoltage : Bool;
      statGetFrame : Struct
         frame0 : Bool;
         frame1 : Bool;
         frame2 : Bool;
         frame21 : Bool;
         frame22 : Bool;
         frame3 : Bool;
         frame31 : Bool;
         frame32 : Bool;
      END_STRUCT;
      statHMI : Struct
         deviceName : String;
         stateCOM : Bool;
         stateDipSwitchTD1 : Bool;
         stateDipSwitchTD2 : Bool;
         stateOutput1 : Int;   // 0=switched-off automatical, no reset possible; 1=switched-off automatical, reset possible; 2= switched-off manual; 3=switched on; 4=defect; 5=device overtemperature; 6=overload; 7=current > nominal value
         stateOutput2 : Int;   // 0=switched-off automatical, no reset possible; 1=switched-off automatical, reset possible; 2= switched-off manual; 3=switched on; 4=defect; 5=device overtemperature; 6=overload; 7=current > nominal value
         stateOutput3 : Int;   // 0=switched-off automatical, no reset possible; 1=switched-off automatical, reset possible; 2= switched-off manual; 3=switched on; 4=defect; 5=device overtemperature; 6=overload; 7=current > nominal value
         stateOutput4 : Int;   // 0=switched-off automatical, no reset possible; 1=switched-off automatical, reset possible; 2= switched-off manual; 3=switched on; 4=defect; 5=device overtemperature; 6=overload; 7=current > nominal value
         stateOutput5 : Int;   // 0=switched-off automatical, no reset possible; 1=switched-off automatical, reset possible; 2= switched-off manual; 3=switched on; 4=defect; 5=device overtemperature; 6=overload; 7=current > nominal value
         stateOutput6 : Int;   // 0=switched-off automatical, no reset possible; 1=switched-off automatical, reset possible; 2= switched-off manual; 3=switched on; 4=defect; 5=device overtemperature; 6=overload; 7=current > nominal value
         stateOutput7 : Int;   // 0=switched-off automatical, no reset possible; 1=switched-off automatical, reset possible; 2= switched-off manual; 3=switched on; 4=defect; 5=device overtemperature; 6=overload; 7=current > nominal value
         stateOutput8 : Int;   // 0=switched-off automatical, no reset possible; 1=switched-off automatical, reset possible; 2= switched-off manual; 3=switched on; 4=defect; 5=device overtemperature; 6=overload; 7=current > nominal value
         outputCurrent1 : Int;   // output current output1
         outputCurrent2 : Int;   // output current output2
         outputCurrent3 : Int;   // output current output3
         outputCurrent4 : Int;   // output current output4
         outputCurrent5 : Int;   // output current output5
         outputCurrent6 : Int;   // output current output6
         outputCurrent7 : Int;   // output current output7
         outputCurrent8 : Int;   // output current output8
         outputCurrentLimit1 : Int;   // output current limit output1
         outputCurrentLimit2 : Int;   // output current limit output2
         outputCurrentLimit3 : Int;   // output current limit output3
         outputCurrentLimit4 : Int;   // output current limit output4
         outputCurrentLimit5 : Int;   // output current limit output5
         outputCurrentLimit6 : Int;   // output current limit output6
         outputCurrentLimit7 : Int;   // output current limit output7
         outputCurrentLimit8 : Int;   // output current limit output8
         reasonOutputSwitchedOff1 : Int;   // 0=output current>limit and output current<1,5xlimit for more than 5sec; 1=current output>1,5xlimit; 2=total overload; 3=Uin<19,4V and output current>limit; 4=Uin<15V; 5=Uin>30V; 6=device overtemperature; 8 to 14=Reserve; 15=default (no automatically switched off)